screen "0030_Tool Allocation" 1280x800, template "Navigation"
   on GenerateScreen: "ToolAllocation_First"()
   Button "Button_1" at 558,753 size 280x42; TextOff '>>>'
      on Press: function_dd21b452("DB939_Tool_alloc_HMI_AllocList_page", 1); "ToolAllocation_First"()
      Visibility <- "DB939_Tool_alloc_HMI_Limit_allocation_list"
   Button "Button_3" at 326,104 size 451x32; TextOff 'Tool Allocation'
   Button "Button_31" at 872,148 size 242x25; TextOff 'Existing Tools'
   Button "Button_35" at 981,96 size 196x42; TextOff 'TOOL Allocation Automatic'; TextList "Tool_Allocation_Mode"
      ProcessValue <- "DB939_Tool_alloc_HMI_Select_hand_automatic_alloc"
      on Press: InvertBit("DB939_Tool_alloc_HMI_Select_hand_automatic_alloc")
   Button "Button_34" at 167,754 size 280x42; TextOff '<<<'
      on Press: function_b9b71300("DB939_Tool_alloc_HMI_AllocList_page", 1); "ToolAllocation_First"()
      Visibility <- "DB939_Tool_alloc_HMI_AllocList_page"
   Button "b_Decress_ToolAllocation" at 272,104 size 46x32; TextOff 'Text'; PictureOff "left arrow"
      on Click: function_b9b71300("DB939_Tool_alloc_HMI_MH_No_selected", 1); "ToolAllocation_Sec"()
      Visibility <- "DB939_Tool_alloc_HMI_Select_hand_automatic_alloc"
   Button "Button_36" at 432,154 size 34x31; TextOff 'Text'; PictureOff "Tongsampah_1"
      Visibility <- "DB939_Tool_alloc_HMI_Alloc_stationTool{1}"
      on Press: SetTag("DB939_Tool_alloc_HMI_Delete_selected_tool", 1)
   Button "Button_37" at 432,194 size 34x31; TextOff 'Text'; PictureOff "Tongsampah_1"
      Visibility <- "DB939_Tool_alloc_HMI_Alloc_stationTool{2}"
      on Press: SetTag("DB939_Tool_alloc_HMI_Delete_selected_tool", 2)
   Button "Button_38" at 432,234 size 34x31; TextOff 'Text'; PictureOff "Tongsampah_1"
      Visibility <- "DB939_Tool_alloc_HMI_Alloc_stationTool{3}"
      on Press: SetTag("DB939_Tool_alloc_HMI_Delete_selected_tool", 3)
   Button "Button_39" at 432,274 size 34x31; TextOff 'Text'; PictureOff "Tongsampah_1"
      Visibility <- "DB939_Tool_alloc_HMI_Alloc_stationTool{4}"
      on Press: SetTag("DB939_Tool_alloc_HMI_Delete_selected_tool", 4)
   Button "Button_40" at 432,314 size 34x31; TextOff 'Text'; PictureOff "Tongsampah_1"
      Visibility <- "DB939_Tool_alloc_HMI_Alloc_stationTool{5}"
      on Press: SetTag("DB939_Tool_alloc_HMI_Delete_selected_tool", 5)
   Button "Button_41" at 432,354 size 34x31; TextOff 'Text'; PictureOff "Tongsampah_1"
      Visibility <- "DB939_Tool_alloc_HMI_Alloc_stationTool{6}"
      on Press: SetTag("DB939_Tool_alloc_HMI_Delete_selected_tool", 6)
   Button "Button_42" at 432,394 size 34x31; TextOff 'Text'; PictureOff "Tongsampah_1"
      Visibility <- "DB939_Tool_alloc_HMI_Alloc_stationTool{7}"
      on Press: SetTag("DB939_Tool_alloc_HMI_Delete_selected_tool", 7)
   Button "Button_43" at 432,434 size 34x31; TextOff 'Text'; PictureOff "Tongsampah_1"
      Visibility <- "DB939_Tool_alloc_HMI_Alloc_stationTool{8}"
      on Press: SetTag("DB939_Tool_alloc_HMI_Delete_selected_tool", 8)
   Button "Button_44" at 432,474 size 34x31; TextOff 'Text'; PictureOff "Tongsampah_1"
      Visibility <- "DB939_Tool_alloc_HMI_Alloc_stationTool{9}"
      on Press: SetTag("DB939_Tool_alloc_HMI_Delete_selected_tool", 9)
   Button "Button_45" at 432,514 size 34x31; TextOff 'Text'; PictureOff "Tongsampah_1"
      Visibility <- "DB939_Tool_alloc_HMI_Alloc_stationTool{10}"
      on Press: SetTag("DB939_Tool_alloc_HMI_Delete_selected_tool", 10)
   Button "Button_46" at 432,554 size 34x31; TextOff 'Text'; PictureOff "Tongsampah_1"
      Visibility <- "DB939_Tool_alloc_HMI_Alloc_stationTool{11}"
      on Press: SetTag("DB939_Tool_alloc_HMI_Delete_selected_tool", 11)
   Button "Button_47" at 432,594 size 34x31; TextOff 'Text'; PictureOff "Tongsampah_1"
      Visibility <- "DB939_Tool_alloc_HMI_Alloc_stationTool{12}"
      on Press: SetTag("DB939_Tool_alloc_HMI_Delete_selected_tool", 12)
   Button "Button_48" at 432,634 size 34x31; TextOff 'Text'; PictureOff "Tongsampah_1"
      Visibility <- "DB939_Tool_alloc_HMI_Alloc_stationTool{13}"
      on Press: SetTag("DB939_Tool_alloc_HMI_Delete_selected_tool", 13)
   Button "Button_49" at 432,674 size 34x31; TextOff 'Text'; PictureOff "Tongsampah_1"
      Visibility <- "DB939_Tool_alloc_HMI_Alloc_stationTool{14}"
      on Press: SetTag("DB939_Tool_alloc_HMI_Delete_selected_tool", 14)
   Button "Button_50" at 432,714 size 34x31; TextOff 'Text'; PictureOff "Tongsampah_1"
      Visibility <- "DB939_Tool_alloc_HMI_Alloc_stationTool{15}"
      on Press: SetTag("DB939_Tool_alloc_HMI_Delete_selected_tool", 15)
   Button "Button_51" at 807,154 size 34x31; TextOff 'Text'; PictureOff "Tongsampah_1"
      Visibility <- "DB939_Tool_alloc_HMI_Alloc_stationTool{16}"
      on Press: SetTag("DB939_Tool_alloc_HMI_Delete_selected_tool", 16)
   Button "Button_52" at 807,194 size 34x31; TextOff 'Text'; PictureOff "Tongsampah_1"
      Visibility <- "DB939_Tool_alloc_HMI_Alloc_stationTool{17}"
      on Press: SetTag("DB939_Tool_alloc_HMI_Delete_selected_tool", 17)
   Button "Button_53" at 807,234 size 34x31; TextOff 'Text'; PictureOff "Tongsampah_1"
      Visibility <- "DB939_Tool_alloc_HMI_Alloc_stationTool{18}"
      on Press: SetTag("DB939_Tool_alloc_HMI_Delete_selected_tool", 18)
   Button "Button_54" at 807,274 size 34x31; TextOff 'Text'; PictureOff "Tongsampah_1"
      Visibility <- "DB939_Tool_alloc_HMI_Alloc_stationTool{19}"
      on Press: SetTag("DB939_Tool_alloc_HMI_Delete_selected_tool", 19)
   Button "Button_55" at 807,314 size 34x31; TextOff 'Text'; PictureOff "Tongsampah_1"
      Visibility <- "DB939_Tool_alloc_HMI_Alloc_stationTool{20}"
      on Press: SetTag("DB939_Tool_alloc_HMI_Delete_selected_tool", 20)
   Button "Button_56" at 807,354 size 34x31; TextOff 'Text'; PictureOff "Tongsampah_1"
      Visibility <- "DB939_Tool_alloc_HMI_Alloc_stationTool{21}"
      on Press: SetTag("DB939_Tool_alloc_HMI_Delete_selected_tool", 21)
   Button "Button_57" at 807,394 size 34x31; TextOff 'Text'; PictureOff "Tongsampah_1"
      Visibility <- "DB939_Tool_alloc_HMI_Alloc_stationTool{22}"
      on Press: SetTag("DB939_Tool_alloc_HMI_Delete_selected_tool", 22)
   Button "Button_58" at 807,434 size 34x31; TextOff 'Text'; PictureOff "Tongsampah_1"
      Visibility <- "DB939_Tool_alloc_HMI_Alloc_stationTool{23}"
      on Press: SetTag("DB939_Tool_alloc_HMI_Delete_selected_tool", 23)
   Button "Button_59" at 807,474 size 34x31; TextOff 'Text'; PictureOff "Tongsampah_1"
      Visibility <- "DB939_Tool_alloc_HMI_Alloc_stationTool{24}"
      on Press: SetTag("DB939_Tool_alloc_HMI_Delete_selected_tool", 24)
   Button "Button_60" at 807,514 size 34x31; TextOff 'Text'; PictureOff "Tongsampah_1"
      Visibility <- "DB939_Tool_alloc_HMI_Alloc_stationTool{25}"
      on Press: SetTag("DB939_Tool_alloc_HMI_Delete_selected_tool", 25)
   Button "Button_61" at 807,554 size 34x31; TextOff 'Text'; PictureOff "Tongsampah_1"
      Visibility <- "DB939_Tool_alloc_HMI_Alloc_stationTool{26}"
      on Press: SetTag("DB939_Tool_alloc_HMI_Delete_selected_tool", 26)
   Button "Button_62" at 807,594 size 34x31; TextOff 'Text'; PictureOff "Tongsampah_1"
      Visibility <- "DB939_Tool_alloc_HMI_Alloc_stationTool{27}"
      on Press: SetTag("DB939_Tool_alloc_HMI_Delete_selected_tool", 27)
   Button "Button_63" at 807,634 size 34x31; TextOff 'Text'; PictureOff "Tongsampah_1"
      Visibility <- "DB939_Tool_alloc_HMI_Alloc_stationTool{28}"
      on Press: SetTag("DB939_Tool_alloc_HMI_Delete_selected_tool", 28)
   Button "Button_64" at 807,674 size 34x31; TextOff 'Text'; PictureOff "Tongsampah_1"
      Visibility <- "DB939_Tool_alloc_HMI_Alloc_stationTool{29}"
      on Press: SetTag("DB939_Tool_alloc_HMI_Delete_selected_tool", 29)
   Button "Button_65" at 807,714 size 34x31; TextOff 'Text'; PictureOff "Tongsampah_1"
      Visibility <- "DB939_Tool_alloc_HMI_Alloc_stationTool{30}"
      on Press: SetTag("DB939_Tool_alloc_HMI_Delete_selected_tool", 30)
   IOField "I/O field_63" at 971,176 size 144x28; FormatPattern ????????????????????
      ProcessValue <- "DB939_Tool_alloc_HMI_SaveSortProg_name{1}"
      Visibility <- "DB939_Tool_alloc_HMI_SaveSortProgs{1}"
   IOField "I/O field_64" at 971,203 size 144x28; FormatPattern ????????????????????
      ProcessValue <- "DB939_Tool_alloc_HMI_SaveSortProg_name{2}"
      Visibility <- "DB939_Tool_alloc_HMI_SaveSortProgs{2}"
   IOField "I/O field_65" at 971,230 size 144x28; FormatPattern ????????????????????
      ProcessValue <- "DB939_Tool_alloc_HMI_SaveSortProg_name{3}"
      Visibility <- "DB939_Tool_alloc_HMI_SaveSortProgs{3}"
   IOField "I/O field_66" at 971,257 size 144x28; FormatPattern ????????????????????
      ProcessValue <- "DB939_Tool_alloc_HMI_SaveSortProg_name{4}"
      Visibility <- "DB939_Tool_alloc_HMI_SaveSortProgs{4}"
   IOField "I/O field_67" at 971,284 size 144x28; FormatPattern ????????????????????
      ProcessValue <- "DB939_Tool_alloc_HMI_SaveSortProg_name{5}"
      Visibility <- "DB939_Tool_alloc_HMI_SaveSortProgs{5}"
   IOField "I/O field_68" at 971,311 size 144x28; FormatPattern ????????????????????
      ProcessValue <- "DB939_Tool_alloc_HMI_SaveSortProg_name{6}"
      Visibility <- "DB939_Tool_alloc_HMI_SaveSortProgs{6}"
   IOField "I/O field_69" at 971,338 size 144x28; FormatPattern ????????????????????
      ProcessValue <- "DB939_Tool_alloc_HMI_SaveSortProg_name{7}"
      Visibility <- "DB939_Tool_alloc_HMI_SaveSortProgs{7}"
   IOField "I/O field_70" at 971,365 size 144x28; FormatPattern ????????????????????
      ProcessValue <- "DB939_Tool_alloc_HMI_SaveSortProg_name{8}"
      Visibility <- "DB939_Tool_alloc_HMI_SaveSortProgs{8}"
   IOField "I/O field_71" at 971,392 size 144x28; FormatPattern ????????????????????
      ProcessValue <- "DB939_Tool_alloc_HMI_SaveSortProg_name{9}"
      Visibility <- "DB939_Tool_alloc_HMI_SaveSortProgs{9}"
   IOField "I/O field_72" at 971,419 size 144x28; FormatPattern ????????????????????
      ProcessValue <- "DB939_Tool_alloc_HMI_SaveSortProg_name{10}"
      Visibility <- "DB939_Tool_alloc_HMI_SaveSortProgs{10}"
   IOField "I/O field_73" at 971,446 size 144x28; FormatPattern ????????????????????
      ProcessValue <- "DB939_Tool_alloc_HMI_SaveSortProg_name{11}"
      Visibility <- "DB939_Tool_alloc_HMI_SaveSortProgs{11}"
   IOField "I/O field_74" at 971,473 size 144x28; FormatPattern ????????????????????
      ProcessValue <- "DB939_Tool_alloc_HMI_SaveSortProg_name{12}"
      Visibility <- "DB939_Tool_alloc_HMI_SaveSortProgs{12}"
   IOField "I/O field_75" at 971,500 size 144x28; FormatPattern ????????????????????
      ProcessValue <- "DB939_Tool_alloc_HMI_SaveSortProg_name{13}"
      Visibility <- "DB939_Tool_alloc_HMI_SaveSortProgs{13}"
   IOField "I/O field_76" at 971,527 size 144x28; FormatPattern ????????????????????
      ProcessValue <- "DB939_Tool_alloc_HMI_SaveSortProg_name{14}"
      Visibility <- "DB939_Tool_alloc_HMI_SaveSortProgs{14}"
   IOField "I/O field_77" at 971,554 size 144x28; FormatPattern ????????????????????
      ProcessValue <- "DB939_Tool_alloc_HMI_SaveSortProg_name{15}"
      Visibility <- "DB939_Tool_alloc_HMI_SaveSortProgs{15}"
   IOField "I/O field_78" at 971,581 size 144x28; FormatPattern ????????????????????
      ProcessValue <- "DB939_Tool_alloc_HMI_SaveSortProg_name{16}"
      Visibility <- "DB939_Tool_alloc_HMI_SaveSortProgs{16}"
   IOField "I/O field_79" at 971,608 size 144x28; FormatPattern ????????????????????
      ProcessValue <- "DB939_Tool_alloc_HMI_SaveSortProg_name{17}"
      Visibility <- "DB939_Tool_alloc_HMI_SaveSortProgs{17}"
   IOField "I/O field_80" at 971,635 size 144x28; FormatPattern ????????????????????
      ProcessValue <- "DB939_Tool_alloc_HMI_SaveSortProg_name{18}"
      Visibility <- "DB939_Tool_alloc_HMI_SaveSortProgs{18}"
   IOField "I/O field_81" at 971,662 size 144x28; FormatPattern ????????????????????
      ProcessValue <- "DB939_Tool_alloc_HMI_SaveSortProg_name{19}"
      Visibility <- "DB939_Tool_alloc_HMI_SaveSortProgs{19}"
   IOField "I/O field_82" at 971,689 size 144x28; FormatPattern ????????????????????
      ProcessValue <- "DB939_Tool_alloc_HMI_SaveSortProg_name{20}"
      Visibility <- "DB939_Tool_alloc_HMI_SaveSortProgs{20}"
   IOField "I/O field_83" at 877,176 size 96x28; FormatPattern 9999
      ProcessValue <- "DB939_Tool_alloc_HMI_SaveSortProgs{1}"
      Visibility <- "DB939_Tool_alloc_HMI_SaveSortProgs{1}"
   IOField "I/O field_84" at 877,203 size 96x28; FormatPattern 9999
      ProcessValue <- "DB939_Tool_alloc_HMI_SaveSortProgs{2}"
      Visibility <- "DB939_Tool_alloc_HMI_SaveSortProgs{2}"
   IOField "I/O field_85" at 877,230 size 96x28; FormatPattern 9999
      ProcessValue <- "DB939_Tool_alloc_HMI_SaveSortProgs{3}"
      Visibility <- "DB939_Tool_alloc_HMI_SaveSortProgs{3}"
   IOField "I/O field_86" at 877,257 size 96x28; FormatPattern 9999
      ProcessValue <- "DB939_Tool_alloc_HMI_SaveSortProgs{4}"
      Visibility <- "DB939_Tool_alloc_HMI_SaveSortProgs{4}"
   IOField "I/O field_87" at 877,284 size 96x28; FormatPattern 9999
      ProcessValue <- "DB939_Tool_alloc_HMI_SaveSortProgs{5}"
      Visibility <- "DB939_Tool_alloc_HMI_SaveSortProgs{5}"
   IOField "I/O field_88" at 877,311 size 96x28; FormatPattern 9999
      ProcessValue <- "DB939_Tool_alloc_HMI_SaveSortProgs{6}"
      Visibility <- "DB939_Tool_alloc_HMI_SaveSortProgs{6}"
   IOField "I/O field_89" at 877,338 size 96x28; FormatPattern 9999
      ProcessValue <- "DB939_Tool_alloc_HMI_SaveSortProgs{7}"
      Visibility <- "DB939_Tool_alloc_HMI_SaveSortProgs{7}"
   IOField "I/O field_90" at 877,365 size 96x28; FormatPattern 9999
      ProcessValue <- "DB939_Tool_alloc_HMI_SaveSortProgs{8}"
      Visibility <- "DB939_Tool_alloc_HMI_SaveSortProgs{8}"
   IOField "I/O field_91" at 877,392 size 96x28; FormatPattern 9999
      ProcessValue <- "DB939_Tool_alloc_HMI_SaveSortProgs{9}"
      Visibility <- "DB939_Tool_alloc_HMI_SaveSortProgs{9}"
   IOField "I/O field_92" at 877,419 size 96x28; FormatPattern 9999
      ProcessValue <- "DB939_Tool_alloc_HMI_SaveSortProgs{10}"
      Visibility <- "DB939_Tool_alloc_HMI_SaveSortProgs{10}"
   IOField "I/O field_93" at 877,446 size 96x28; FormatPattern 9999
      ProcessValue <- "DB939_Tool_alloc_HMI_SaveSortProgs{11}"
      Visibility <- "DB939_Tool_alloc_HMI_SaveSortProgs{11}"
   IOField "I/O field_94" at 877,473 size 96x28; FormatPattern 9999
      ProcessValue <- "DB939_Tool_alloc_HMI_SaveSortProgs{12}"
      Visibility <- "DB939_Tool_alloc_HMI_SaveSortProgs{12}"
   IOField "I/O field_95" at 877,500 size 96x28; FormatPattern 9999
      ProcessValue <- "DB939_Tool_alloc_HMI_SaveSortProgs{13}"
      Visibility <- "DB939_Tool_alloc_HMI_SaveSortProgs{13}"
   IOField "I/O field_96" at 877,527 size 96x28; FormatPattern 9999
      ProcessValue <- "DB939_Tool_alloc_HMI_SaveSortProgs{14}"
      Visibility <- "DB939_Tool_alloc_HMI_SaveSortProgs{14}"
   IOField "I/O field_97" at 877,554 size 96x28; FormatPattern 9999
      ProcessValue <- "DB939_Tool_alloc_HMI_SaveSortProgs{15}"
      Visibility <- "DB939_Tool_alloc_HMI_SaveSortProgs{15}"
   IOField "I/O field_98" at 877,581 size 96x28; FormatPattern 9999
      ProcessValue <- "DB939_Tool_alloc_HMI_SaveSortProgs{16}"
      Visibility <- "DB939_Tool_alloc_HMI_SaveSortProgs{16}"
   IOField "I/O field_99" at 877,608 size 96x28; FormatPattern 9999
      ProcessValue <- "DB939_Tool_alloc_HMI_SaveSortProgs{17}"
      Visibility <- "DB939_Tool_alloc_HMI_SaveSortProgs{17}"
   IOField "I/O field_100" at 877,635 size 96x28; FormatPattern 9999
      ProcessValue <- "DB939_Tool_alloc_HMI_SaveSortProgs{18}"
      Visibility <- "DB939_Tool_alloc_HMI_SaveSortProgs{18}"
   IOField "I/O field_101" at 877,662 size 96x28; FormatPattern 9999
      ProcessValue <- "DB939_Tool_alloc_HMI_SaveSortProgs{19}"
      Visibility <- "DB939_Tool_alloc_HMI_SaveSortProgs{19}"
   IOField "I/O field_102" at 877,689 size 96x28; FormatPattern 9999
      ProcessValue <- "DB939_Tool_alloc_HMI_SaveSortProgs{20}"
      Visibility <- "DB939_Tool_alloc_HMI_SaveSortProgs{20}"
   Button "Button_66" at 1128,183 size 42x224; TextOff '˄˄˄'
      on Press: SetBit("DB939_Tool_alloc_HMI_SavedProgs_increase")
      Visibility <- "DB939_Tool_alloc_HMI_SavedProgs_increase_visible"
   Button "Button_67" at 1128,485 size 42x224; TextOff 'VVV'
      on Press: SetBit("DB939_Tool_alloc_HMI_SavedProgs_decrease")
      Visibility <- "DB939_Tool_alloc_HMI_SavedProgs_decrease_visible"
   Button "b_Incress_ToolAllocation" at 786,104 size 46x32; TextOff 'Text'; PictureOff "right arrow"
      on Click: function_dd21b452("DB939_Tool_alloc_HMI_MH_No_selected", 1); "ToolAllocation_Sec"()
      Visibility <- "DB939_Tool_alloc_HMI_Select_hand_automatic_alloc"
   IOField "I/O field_5" at 179,152 size 73x35; Authorization "User administration"; FormatPattern 999
      ProcessValue <- "DB939_Tool_alloc_HMI_Alloc_stationTool{1}"
      Visibility <- "DB939_Tool_alloc_HMI_Limit_allocation_list"
      Appearance <- "DB939_Tool_alloc_HMI_Selected_prog"
   Button "Button_6" at 123,152 size 50x35; TextOff '.'
      Visibility <- "DB939_Tool_alloc_HMI_Limit_allocation_list"
      on Press: SetTag("DB939_Tool_alloc_HMI_Selected_prog", 1)
      Appearance <- "DB939_Tool_alloc_HMI_Selected_prog"
   Button "Button_2" at 123,192 size 50x35; TextOff '.'
      Visibility <- "DB939_Tool_alloc_HMI_Limit_allocation_list"
      on Press: SetTag("DB939_Tool_alloc_HMI_Selected_prog", 2)
      Appearance <- "DB939_Tool_alloc_HMI_Selected_prog"
   Button "Button_4" at 123,232 size 50x35; TextOff '.'
      Visibility <- "DB939_Tool_alloc_HMI_Limit_allocation_list"
      on Press: SetTag("DB939_Tool_alloc_HMI_Selected_prog", 3)
      Appearance <- "DB939_Tool_alloc_HMI_Selected_prog"
   Button "Button_5" at 123,272 size 50x35; TextOff '.'
      Visibility <- "DB939_Tool_alloc_HMI_Limit_allocation_list"
      on Press: SetTag("DB939_Tool_alloc_HMI_Selected_prog", 4)
      Appearance <- "DB939_Tool_alloc_HMI_Selected_prog"
   Button "Button_7" at 123,312 size 50x35; TextOff '.'
      Visibility <- "DB939_Tool_alloc_HMI_Limit_allocation_list"
      on Press: SetTag("DB939_Tool_alloc_HMI_Selected_prog", 5)
      Appearance <- "DB939_Tool_alloc_HMI_Selected_prog"
   Button "Button_8" at 123,352 size 50x35; TextOff '.'
      Visibility <- "DB939_Tool_alloc_HMI_Limit_allocation_list"
      on Press: SetTag("DB939_Tool_alloc_HMI_Selected_prog", 6)
      Appearance <- "DB939_Tool_alloc_HMI_Selected_prog"
   Button "Button_9" at 123,392 size 50x35; TextOff '.'
      Visibility <- "DB939_Tool_alloc_HMI_Limit_allocation_list"
      on Press: SetTag("DB939_Tool_alloc_HMI_Selected_prog", 7)
      Appearance <- "DB939_Tool_alloc_HMI_Selected_prog"
   Button "Button_10" at 123,432 size 50x35; TextOff '.'
      on Press: SetTag("DB939_Tool_alloc_HMI_Selected_prog", 8)
      Appearance <- "DB939_Tool_alloc_HMI_Selected_prog"
      Visibility <- "DB939_Tool_alloc_HMI_Limit_allocation_list"
   Button "Button_11" at 123,472 size 50x35; TextOff '.'
      Visibility <- "DB939_Tool_alloc_HMI_Limit_allocation_list"
      on Press: SetTag("DB939_Tool_alloc_HMI_Selected_prog", 9)
      Appearance <- "DB939_Tool_alloc_HMI_Selected_prog"
   Button "Button_12" at 123,512 size 50x35; TextOff '.'
      Visibility <- "DB939_Tool_alloc_HMI_Limit_allocation_list"
      on Press: SetTag("DB939_Tool_alloc_HMI_Selected_prog", 10)
      Appearance <- "DB939_Tool_alloc_HMI_Selected_prog"
   Button "Button_13" at 123,552 size 50x35; TextOff '.'
      Visibility <- "DB939_Tool_alloc_HMI_Limit_allocation_list"
      on Press: SetTag("DB939_Tool_alloc_HMI_Selected_prog", 11)
      Appearance <- "DB939_Tool_alloc_HMI_Selected_prog"
   Button "Button_14" at 123,592 size 50x35; TextOff '.'
      Visibility <- "DB939_Tool_alloc_HMI_Limit_allocation_list"
      on Press: SetTag("DB939_Tool_alloc_HMI_Selected_prog", 12)
      Appearance <- "DB939_Tool_alloc_HMI_Selected_prog"
   Button "Button_15" at 123,632 size 50x35; TextOff '.'
      Visibility <- "DB939_Tool_alloc_HMI_Limit_allocation_list"
      on Press: SetTag("DB939_Tool_alloc_HMI_Selected_prog", 13)
      Appearance <- "DB939_Tool_alloc_HMI_Selected_prog"
   Button "Button_16" at 123,672 size 50x35; TextOff '.'
      Visibility <- "DB939_Tool_alloc_HMI_Limit_allocation_list"
      on Press: SetTag("DB939_Tool_alloc_HMI_Selected_prog", 14)
      Appearance <- "DB939_Tool_alloc_HMI_Selected_prog"
   Button "Button_17" at 496,152 size 50x35; TextOff '.'
      Visibility <- "DB939_Tool_alloc_HMI_Limit_allocation_list"
      on Press: SetTag("DB939_Tool_alloc_HMI_Selected_prog", 16)
      Appearance <- "DB939_Tool_alloc_HMI_Selected_prog"
   Button "Button_18" at 496,192 size 50x35; TextOff '.'
      Visibility <- "DB939_Tool_alloc_HMI_Limit_allocation_list"
      on Press: SetTag("DB939_Tool_alloc_HMI_Selected_prog", 17)
      Appearance <- "DB939_Tool_alloc_HMI_Selected_prog"
   Button "Button_19" at 496,232 size 50x35; TextOff '.'
      Visibility <- "DB939_Tool_alloc_HMI_Limit_allocation_list"
      on Press: SetTag("DB939_Tool_alloc_HMI_Selected_prog", 18)
      Appearance <- "DB939_Tool_alloc_HMI_Selected_prog"
   Button "Button_20" at 496,272 size 50x35; TextOff '.'
      Visibility <- "DB939_Tool_alloc_HMI_Limit_allocation_list"
      on Press: SetTag("DB939_Tool_alloc_HMI_Selected_prog", 19)
      Appearance <- "DB939_Tool_alloc_HMI_Selected_prog"
   Button "Button_21" at 496,312 size 50x35; TextOff '.'
      Visibility <- "DB939_Tool_alloc_HMI_Limit_allocation_list"
      on Press: SetTag("DB939_Tool_alloc_HMI_Selected_prog", 20)
      Appearance <- "DB939_Tool_alloc_HMI_Selected_prog"
   Button "Button_22" at 496,352 size 50x35; TextOff '.'
      Visibility <- "DB939_Tool_alloc_HMI_Limit_allocation_list"
      on Press: SetTag("DB939_Tool_alloc_HMI_Selected_prog", 21)
      Appearance <- "DB939_Tool_alloc_HMI_Selected_prog"
   Button "Button_23" at 496,392 size 50x35; TextOff '.'
      Visibility <- "DB939_Tool_alloc_HMI_Limit_allocation_list"
      on Press: SetTag("DB939_Tool_alloc_HMI_Selected_prog", 22)
      Appearance <- "DB939_Tool_alloc_HMI_Selected_prog"
   Button "Button_24" at 496,432 size 50x35; TextOff '.'
      Visibility <- "DB939_Tool_alloc_HMI_Limit_allocation_list"
      on Press: SetTag("DB939_Tool_alloc_HMI_Selected_prog", 23)
      Appearance <- "DB939_Tool_alloc_HMI_Selected_prog"
   Button "Button_25" at 496,472 size 50x35; TextOff 'Text'
      Visibility <- "DB939_Tool_alloc_HMI_Limit_allocation_list"
      on Press: SetTag("DB939_Tool_alloc_HMI_Selected_prog", 24)
      Appearance <- "DB939_Tool_alloc_HMI_Selected_prog"
   Button "Button_26" at 496,512 size 50x35; TextOff 'Text'
      Visibility <- "DB939_Tool_alloc_HMI_Limit_allocation_list"
      on Press: SetTag("DB939_Tool_alloc_HMI_Selected_prog", 25)
      Appearance <- "DB939_Tool_alloc_HMI_Selected_prog"
   Button "Button_27" at 496,552 size 50x35; TextOff '.'
      Visibility <- "DB939_Tool_alloc_HMI_Limit_allocation_list"
      on Press: SetTag("DB939_Tool_alloc_HMI_Selected_prog", 26)
      Appearance <- "DB939_Tool_alloc_HMI_Selected_prog"
   Button "Button_28" at 496,592 size 50x35; TextOff '.'
      Visibility <- "DB939_Tool_alloc_HMI_Limit_allocation_list"
      on Press: SetTag("DB939_Tool_alloc_HMI_Selected_prog", 27)
      Appearance <- "DB939_Tool_alloc_HMI_Selected_prog"
   Button "Button_29" at 496,632 size 50x35; TextOff '.'
      Visibility <- "DB939_Tool_alloc_HMI_Limit_allocation_list"
      on Press: SetTag("DB939_Tool_alloc_HMI_Selected_prog", 28)
      Appearance <- "DB939_Tool_alloc_HMI_Selected_prog"
   Button "Button_30" at 496,672 size 50x35; TextOff '.'
      Visibility <- "DB939_Tool_alloc_HMI_Limit_allocation_list"
      on Press: SetTag("DB939_Tool_alloc_HMI_Selected_prog", 29)
      Appearance <- "DB939_Tool_alloc_HMI_Selected_prog"
   IOField "Station_Tool_2" at 179,192 size 73x35; Authorization "User administration"; FormatPattern 999
      ProcessValue <- "DB939_Tool_alloc_HMI_Alloc_stationTool{2}"
      Visibility <- "DB939_Tool_alloc_HMI_Limit_allocation_list"
      Appearance <- "DB939_Tool_alloc_HMI_Selected_prog"
   IOField "I/O field_2" at 179,232 size 73x35; Authorization "User administration"; FormatPattern 999
      ProcessValue <- "DB939_Tool_alloc_HMI_Alloc_stationTool{3}"
      Visibility <- "DB939_Tool_alloc_HMI_Limit_allocation_list"
      Appearance <- "DB939_Tool_alloc_HMI_Selected_prog"
   IOField "I/O field_3" at 179,272 size 73x35; Authorization "User administration"; FormatPattern 999
      ProcessValue <- "DB939_Tool_alloc_HMI_Alloc_stationTool{4}"
      Visibility <- "DB939_Tool_alloc_HMI_Limit_allocation_list"
      Appearance <- "DB939_Tool_alloc_HMI_Selected_prog"
   IOField "I/O field_4" at 179,312 size 73x35; Authorization "User administration"; FormatPattern 999
      ProcessValue <- "DB939_Tool_alloc_HMI_Alloc_stationTool{5}"
      Visibility <- "DB939_Tool_alloc_HMI_Limit_allocation_list"
      Appearance <- "DB939_Tool_alloc_HMI_Selected_prog"
   IOField "I/O field_6" at 179,352 size 73x35; Authorization "User administration"; FormatPattern 999
      ProcessValue <- "DB939_Tool_alloc_HMI_Alloc_stationTool{6}"
      Visibility <- "DB939_Tool_alloc_HMI_Limit_allocation_list"
      Appearance <- "DB939_Tool_alloc_HMI_Selected_prog"
   IOField "I/O field_7" at 179,392 size 73x35; Authorization "User administration"; FormatPattern 999
      ProcessValue <- "DB939_Tool_alloc_HMI_Alloc_stationTool{7}"
      Visibility <- "DB939_Tool_alloc_HMI_Limit_allocation_list"
      Appearance <- "DB939_Tool_alloc_HMI_Selected_prog"
   IOField "I/O field_8" at 179,432 size 73x35; Authorization "User administration"; FormatPattern 999
      ProcessValue <- "DB939_Tool_alloc_HMI_Alloc_stationTool{8}"
      Appearance <- "DB939_Tool_alloc_HMI_Selected_prog"
      Visibility <- "DB939_Tool_alloc_HMI_Limit_allocation_list"
   IOField "I/O field_9" at 179,472 size 73x35; Authorization "User administration"; FormatPattern 999
      ProcessValue <- "DB939_Tool_alloc_HMI_Alloc_stationTool{9}"
      Visibility <- "DB939_Tool_alloc_HMI_Limit_allocation_list"
      Appearance <- "DB939_Tool_alloc_HMI_Selected_prog"
   IOField "I/O field_10" at 179,512 size 73x35; Authorization "User administration"; FormatPattern 999
      ProcessValue <- "DB939_Tool_alloc_HMI_Alloc_stationTool{10}"
      Visibility <- "DB939_Tool_alloc_HMI_Limit_allocation_list"
      Appearance <- "DB939_Tool_alloc_HMI_Selected_prog"
   IOField "I/O field_11" at 179,552 size 73x35; Authorization "User administration"; FormatPattern 999
      ProcessValue <- "DB939_Tool_alloc_HMI_Alloc_stationTool{11}"
      Visibility <- "DB939_Tool_alloc_HMI_Limit_allocation_list"
      Appearance <- "DB939_Tool_alloc_HMI_Selected_prog"
   IOField "I/O field_12" at 179,592 size 73x35; Authorization "User administration"; FormatPattern 999
      ProcessValue <- "DB939_Tool_alloc_HMI_Alloc_stationTool{12}"
      Visibility <- "DB939_Tool_alloc_HMI_Limit_allocation_list"
      Appearance <- "DB939_Tool_alloc_HMI_Selected_prog"
   IOField "I/O field_13" at 179,632 size 73x35; Authorization "User administration"; FormatPattern 999
      ProcessValue <- "DB939_Tool_alloc_HMI_Alloc_stationTool{13}"
      Visibility <- "DB939_Tool_alloc_HMI_Limit_allocation_list"
      Appearance <- "DB939_Tool_alloc_HMI_Selected_prog"
   IOField "I/O field_14" at 179,672 size 73x35; Authorization "User administration"; FormatPattern 999
      ProcessValue <- "DB939_Tool_alloc_HMI_Alloc_stationTool{14}"
      Visibility <- "DB939_Tool_alloc_HMI_Limit_allocation_list"
      Appearance <- "DB939_Tool_alloc_HMI_Selected_prog"
   IOField "I/O field_15" at 552,152 size 73x35; Authorization "User administration"; FormatPattern 999
      ProcessValue <- "DB939_Tool_alloc_HMI_Alloc_stationTool{16}"
      Visibility <- "DB939_Tool_alloc_HMI_Limit_allocation_list"
      Appearance <- "DB939_Tool_alloc_HMI_Selected_prog"
   IOField "I/O field_16" at 552,192 size 73x35; Authorization "User administration"; FormatPattern 999
      ProcessValue <- "DB939_Tool_alloc_HMI_Alloc_stationTool{17}"
      Visibility <- "DB939_Tool_alloc_HMI_Limit_allocation_list"
      Appearance <- "DB939_Tool_alloc_HMI_Selected_prog"
   IOField "I/O field_17" at 552,232 size 73x35; Authorization "User administration"; FormatPattern 999
      ProcessValue <- "DB939_Tool_alloc_HMI_Alloc_stationTool{18}"
      Visibility <- "DB939_Tool_alloc_HMI_Limit_allocation_list"
      Appearance <- "DB939_Tool_alloc_HMI_Selected_prog"
   IOField "I/O field_18" at 552,272 size 73x35; Authorization "User administration"; FormatPattern 999
      ProcessValue <- "DB939_Tool_alloc_HMI_Alloc_stationTool{19}"
      Visibility <- "DB939_Tool_alloc_HMI_Limit_allocation_list"
      Appearance <- "DB939_Tool_alloc_HMI_Selected_prog"
   IOField "I/O field_19" at 552,312 size 73x35; Authorization "User administration"; FormatPattern 999
      ProcessValue <- "DB939_Tool_alloc_HMI_Alloc_stationTool{20}"
      Visibility <- "DB939_Tool_alloc_HMI_Limit_allocation_list"
      Appearance <- "DB939_Tool_alloc_HMI_Selected_prog"
   IOField "I/O field_20" at 552,352 size 73x35; Authorization "User administration"; FormatPattern 999
      ProcessValue <- "DB939_Tool_alloc_HMI_Alloc_stationTool{21}"
      Visibility <- "DB939_Tool_alloc_HMI_Limit_allocation_list"
      Appearance <- "DB939_Tool_alloc_HMI_Selected_prog"
   IOField "I/O field_21" at 552,392 size 73x35; Authorization "User administration"; FormatPattern 999
      ProcessValue <- "DB939_Tool_alloc_HMI_Alloc_stationTool{22}"
      Visibility <- "DB939_Tool_alloc_HMI_Limit_allocation_list"
      Appearance <- "DB939_Tool_alloc_HMI_Selected_prog"
   IOField "I/O field_22" at 552,432 size 73x35; Authorization "User administration"; FormatPattern 999
      ProcessValue <- "DB939_Tool_alloc_HMI_Alloc_stationTool{23}"
      Visibility <- "DB939_Tool_alloc_HMI_Limit_allocation_list"
      Appearance <- "DB939_Tool_alloc_HMI_Selected_prog"
   IOField "I/O field_23" at 552,472 size 73x35; Authorization "User administration"; FormatPattern 999
      ProcessValue <- "DB939_Tool_alloc_HMI_Alloc_stationTool{24}"
      Visibility <- "DB939_Tool_alloc_HMI_Limit_allocation_list"
      Appearance <- "DB939_Tool_alloc_HMI_Selected_prog"
   IOField "I/O field_24" at 552,512 size 73x35; Authorization "User administration"; FormatPattern 999
      ProcessValue <- "DB939_Tool_alloc_HMI_Alloc_stationTool{25}"
      Visibility <- "DB939_Tool_alloc_HMI_Limit_allocation_list"
      Appearance <- "DB939_Tool_alloc_HMI_Selected_prog"
   IOField "I/O field_25" at 552,552 size 73x35; Authorization "User administration"; FormatPattern 999
      ProcessValue <- "DB939_Tool_alloc_HMI_Alloc_stationTool{26}"
      Visibility <- "DB939_Tool_alloc_HMI_Limit_allocation_list"
      Appearance <- "DB939_Tool_alloc_HMI_Selected_prog"
   IOField "I/O field_26" at 552,592 size 73x35; Authorization "User administration"; FormatPattern 999
      ProcessValue <- "DB939_Tool_alloc_HMI_Alloc_stationTool{27}"
      Visibility <- "DB939_Tool_alloc_HMI_Limit_allocation_list"
      Appearance <- "DB939_Tool_alloc_HMI_Selected_prog"
   IOField "I/O field_27" at 552,632 size 73x35; Authorization "User administration"; FormatPattern 999
      ProcessValue <- "DB939_Tool_alloc_HMI_Alloc_stationTool{28}"
      Visibility <- "DB939_Tool_alloc_HMI_Limit_allocation_list"
      Appearance <- "DB939_Tool_alloc_HMI_Selected_prog"
   IOField "I/O field_28" at 552,672 size 73x35; Authorization "User administration"; FormatPattern 999
      ProcessValue <- "DB939_Tool_alloc_HMI_Alloc_stationTool{29}"
      Visibility <- "DB939_Tool_alloc_HMI_Limit_allocation_list"
      Appearance <- "DB939_Tool_alloc_HMI_Selected_prog"
   IOField "I/O field_29" at 259,152 size 159x35; Authorization "User administration"; FormatPattern ????????????????????
      ProcessValue <- "DB939_Tool_alloc_HMI_Alloc_tool_name{1}"
      Visibility <- "DB939_Tool_alloc_HMI_Limit_allocation_list"
      Appearance <- "DB939_Tool_alloc_HMI_Selected_prog"
   IOField "I/O field_30" at 260,192 size 159x35; Authorization "User administration"; FormatPattern ????????????????????
      ProcessValue <- "DB939_Tool_alloc_HMI_Alloc_tool_name{2}"
      Visibility <- "DB939_Tool_alloc_HMI_Limit_allocation_list"
      Appearance <- "DB939_Tool_alloc_HMI_Selected_prog"
   IOField "I/O field_31" at 260,232 size 159x35; Authorization "User administration"; FormatPattern ????????????????????
      ProcessValue <- "DB939_Tool_alloc_HMI_Alloc_tool_name{3}"
      Visibility <- "DB939_Tool_alloc_HMI_Limit_allocation_list"
      Appearance <- "DB939_Tool_alloc_HMI_Selected_prog"
   IOField "I/O field_32" at 260,272 size 159x35; Authorization "User administration"; FormatPattern ????????????????????
      ProcessValue <- "DB939_Tool_alloc_HMI_Alloc_tool_name{4}"
      Visibility <- "DB939_Tool_alloc_HMI_Limit_allocation_list"
      Appearance <- "DB939_Tool_alloc_HMI_Selected_prog"
   IOField "I/O field_33" at 260,312 size 159x35; Authorization "User administration"; FormatPattern ????????????????????
      ProcessValue <- "DB939_Tool_alloc_HMI_Alloc_tool_name{5}"
      Visibility <- "DB939_Tool_alloc_HMI_Limit_allocation_list"
      Appearance <- "DB939_Tool_alloc_HMI_Selected_prog"
   IOField "I/O field_34" at 260,352 size 159x35; Authorization "User administration"; FormatPattern ????????????????????
      ProcessValue <- "DB939_Tool_alloc_HMI_Alloc_tool_name{6}"
      Visibility <- "DB939_Tool_alloc_HMI_Limit_allocation_list"
      Appearance <- "DB939_Tool_alloc_HMI_Selected_prog"
   IOField "I/O field_35" at 260,392 size 159x35; Authorization "User administration"; FormatPattern ????????????????????
      ProcessValue <- "DB939_Tool_alloc_HMI_Alloc_tool_name{7}"
      Visibility <- "DB939_Tool_alloc_HMI_Limit_allocation_list"
      Appearance <- "DB939_Tool_alloc_HMI_Selected_prog"
   IOField "I/O field_36" at 260,432 size 159x35; Authorization "User administration"; FormatPattern ????????????????????
      ProcessValue <- "DB939_Tool_alloc_HMI_Alloc_tool_name{8}"
      Appearance <- "DB939_Tool_alloc_HMI_Selected_prog"
      Visibility <- "DB939_Tool_alloc_HMI_Limit_allocation_list"
   IOField "I/O field_37" at 260,472 size 159x35; Authorization "User administration"; FormatPattern ????????????????????
      ProcessValue <- "DB939_Tool_alloc_HMI_Alloc_tool_name{9}"
      Visibility <- "DB939_Tool_alloc_HMI_Limit_allocation_list"
      Appearance <- "DB939_Tool_alloc_HMI_Selected_prog"
   IOField "I/O field_38" at 260,512 size 159x35; Authorization "User administration"; FormatPattern ????????????????????
      ProcessValue <- "DB939_Tool_alloc_HMI_Alloc_tool_name{10}"
      Visibility <- "DB939_Tool_alloc_HMI_Limit_allocation_list"
      Appearance <- "DB939_Tool_alloc_HMI_Selected_prog"
   IOField "I/O field_39" at 260,552 size 159x35; Authorization "User administration"; FormatPattern ????????????????????
      ProcessValue <- "DB939_Tool_alloc_HMI_Alloc_tool_name{11}"
      Visibility <- "DB939_Tool_alloc_HMI_Limit_allocation_list"
      Appearance <- "DB939_Tool_alloc_HMI_Selected_prog"
   IOField "I/O field_40" at 260,592 size 159x35; Authorization "User administration"; FormatPattern ????????????????????
      ProcessValue <- "DB939_Tool_alloc_HMI_Alloc_tool_name{12}"
      Visibility <- "DB939_Tool_alloc_HMI_Limit_allocation_list"
      Appearance <- "DB939_Tool_alloc_HMI_Selected_prog"
   IOField "I/O field_41" at 260,632 size 159x35; Authorization "User administration"; FormatPattern ????????????????????
      ProcessValue <- "DB939_Tool_alloc_HMI_Alloc_tool_name{13}"
      Visibility <- "DB939_Tool_alloc_HMI_Limit_allocation_list"
      Appearance <- "DB939_Tool_alloc_HMI_Selected_prog"
   IOField "I/O field_42" at 260,672 size 159x35; Authorization "User administration"; FormatPattern ????????????????????
      ProcessValue <- "DB939_Tool_alloc_HMI_Alloc_tool_name{14}"
      Visibility <- "DB939_Tool_alloc_HMI_Limit_allocation_list"
      Appearance <- "DB939_Tool_alloc_HMI_Selected_prog"
   IOField "I/O field_43" at 632,152 size 159x35; Authorization "User administration"; FormatPattern ????????????????????
      ProcessValue <- "DB939_Tool_alloc_HMI_Alloc_tool_name{16}"
      Visibility <- "DB939_Tool_alloc_HMI_Limit_allocation_list"
      Appearance <- "DB939_Tool_alloc_HMI_Selected_prog"
   IOField "I/O field_44" at 632,192 size 159x35; Authorization "User administration"; FormatPattern ????????????????????
      ProcessValue <- "DB939_Tool_alloc_HMI_Alloc_tool_name{17}"
      Visibility <- "DB939_Tool_alloc_HMI_Limit_allocation_list"
      Appearance <- "DB939_Tool_alloc_HMI_Selected_prog"
   IOField "I/O field_45" at 632,232 size 159x35; Authorization "User administration"; FormatPattern ????????????????????
      ProcessValue <- "DB939_Tool_alloc_HMI_Alloc_tool_name{18}"
      Visibility <- "DB939_Tool_alloc_HMI_Limit_allocation_list"
      Appearance <- "DB939_Tool_alloc_HMI_Selected_prog"
   IOField "I/O field_46" at 632,272 size 159x35; Authorization "User administration"; FormatPattern ????????????????????
      ProcessValue <- "DB939_Tool_alloc_HMI_Alloc_tool_name{19}"
      Visibility <- "DB939_Tool_alloc_HMI_Limit_allocation_list"
      Appearance <- "DB939_Tool_alloc_HMI_Selected_prog"
   IOField "I/O field_47" at 632,312 size 159x35; Authorization "User administration"; FormatPattern ????????????????????
      ProcessValue <- "DB939_Tool_alloc_HMI_Alloc_tool_name{20}"
      Visibility <- "DB939_Tool_alloc_HMI_Limit_allocation_list"
      Appearance <- "DB939_Tool_alloc_HMI_Selected_prog"
   IOField "I/O field_48" at 632,352 size 159x35; Authorization "User administration"; FormatPattern ????????????????????
      ProcessValue <- "DB939_Tool_alloc_HMI_Alloc_tool_name{21}"
      Visibility <- "DB939_Tool_alloc_HMI_Limit_allocation_list"
      Appearance <- "DB939_Tool_alloc_HMI_Selected_prog"
   IOField "I/O field_49" at 632,392 size 159x35; Authorization "User administration"; FormatPattern ????????????????????
      ProcessValue <- "DB939_Tool_alloc_HMI_Alloc_tool_name{22}"
      Visibility <- "DB939_Tool_alloc_HMI_Limit_allocation_list"
      Appearance <- "DB939_Tool_alloc_HMI_Selected_prog"
   IOField "I/O field_50" at 632,432 size 159x35; Authorization "User administration"; FormatPattern ????????????????????
      ProcessValue <- "DB939_Tool_alloc_HMI_Alloc_tool_name{23}"
      Visibility <- "DB939_Tool_alloc_HMI_Limit_allocation_list"
      Appearance <- "DB939_Tool_alloc_HMI_Selected_prog"
   IOField "I/O field_51" at 632,472 size 159x35; Authorization "User administration"; FormatPattern ????????????????????
      ProcessValue <- "DB939_Tool_alloc_HMI_Alloc_tool_name{24}"
      Visibility <- "DB939_Tool_alloc_HMI_Limit_allocation_list"
      Appearance <- "DB939_Tool_alloc_HMI_Selected_prog"
   IOField "I/O field_52" at 632,512 size 159x35; Authorization "User administration"; FormatPattern ????????????????????
      ProcessValue <- "DB939_Tool_alloc_HMI_Alloc_tool_name{25}"
      Visibility <- "DB939_Tool_alloc_HMI_Limit_allocation_list"
      Appearance <- "DB939_Tool_alloc_HMI_Selected_prog"
   IOField "I/O field_53" at 632,552 size 159x35; Authorization "User administration"; FormatPattern ????????????????????
      ProcessValue <- "DB939_Tool_alloc_HMI_Alloc_tool_name{26}"
      Visibility <- "DB939_Tool_alloc_HMI_Limit_allocation_list"
      Appearance <- "DB939_Tool_alloc_HMI_Selected_prog"
   IOField "I/O field_54" at 632,592 size 159x35; Authorization "User administration"; FormatPattern ????????????????????
      ProcessValue <- "DB939_Tool_alloc_HMI_Alloc_tool_name{27}"
      Visibility <- "DB939_Tool_alloc_HMI_Limit_allocation_list"
      Appearance <- "DB939_Tool_alloc_HMI_Selected_prog"
   IOField "I/O field_55" at 632,632 size 159x35; Authorization "User administration"; FormatPattern ????????????????????
      ProcessValue <- "DB939_Tool_alloc_HMI_Alloc_tool_name{28}"
      Visibility <- "DB939_Tool_alloc_HMI_Limit_allocation_list"
      Appearance <- "DB939_Tool_alloc_HMI_Selected_prog"
   IOField "I/O field_56" at 632,672 size 159x35; Authorization "User administration"; FormatPattern ????????????????????
      ProcessValue <- "DB939_Tool_alloc_HMI_Alloc_tool_name{29}"
      Visibility <- "DB939_Tool_alloc_HMI_Limit_allocation_list"
      Appearance <- "DB939_Tool_alloc_HMI_Selected_prog"
   Button "Button_32" at 496,710 size 50x35; TextOff '.'
      Visibility <- "DB939_Tool_alloc_HMI_Limit_allocation_list"
      on Press: SetTag("DB939_Tool_alloc_HMI_Selected_prog", 30)
      Appearance <- "DB939_Tool_alloc_HMI_Selected_prog"
   IOField "I/O field_57" at 551,707 size 73x35; Authorization "User administration"; FormatPattern 999
      ProcessValue <- "DB939_Tool_alloc_HMI_Alloc_stationTool{30}"
      Visibility <- "DB939_Tool_alloc_HMI_Limit_allocation_list"
      Appearance <- "DB939_Tool_alloc_HMI_Selected_prog"
   IOField "I/O field_58" at 631,707 size 159x35; Authorization "User administration"; FormatPattern ????????????????????
      ProcessValue <- "DB939_Tool_alloc_HMI_Alloc_tool_name{30}"
      Visibility <- "DB939_Tool_alloc_HMI_Limit_allocation_list"
      Appearance <- "DB939_Tool_alloc_HMI_Selected_prog"
   Button "Button_33" at 124,713 size 50x35; TextOff '.'
      Visibility <- "DB939_Tool_alloc_HMI_Limit_allocation_list"
      on Press: SetTag("DB939_Tool_alloc_HMI_Selected_prog", 15)
      Appearance <- "DB939_Tool_alloc_HMI_Selected_prog"
   IOField "I/O field_59" at 180,712 size 73x35; Authorization "User administration"; FormatPattern 999
      ProcessValue <- "DB939_Tool_alloc_HMI_Alloc_stationTool{15}"
      Visibility <- "DB939_Tool_alloc_HMI_Limit_allocation_list"
      Appearance <- "DB939_Tool_alloc_HMI_Selected_prog"
   IOField "I/O field_60" at 260,712 size 159x35; Authorization "User administration"; FormatPattern ????????????????????
      ProcessValue <- "DB939_Tool_alloc_HMI_Alloc_tool_name{15}"
      Visibility <- "DB939_Tool_alloc_HMI_Limit_allocation_list"
      Appearance <- "DB939_Tool_alloc_HMI_Selected_prog"
   IOField "I/O field_61" at 465,756 size 73x35; FormatPattern 999
      ProcessValue <- "DB939_Tool_alloc_HMI_AllocList_page"
      Visibility <- "DB939_Tool_alloc_HMI_Limit_allocation_list"
   IOField "I/O field_62" at 734,108 size 39x25; FormatPattern 99
      ProcessValue <- "DB939_Tool_alloc_HMI_MH_No_selected"
      Visibility <- "DB939_Tool_alloc_HMI_Select_hand_automatic_alloc"
   Button "Button_68" at 864,176 size 256x28; TextOff 'Text'
      on Press: SetTag("Tag_1", 1)
      Visibility <- "DB939_Tool_alloc_HMI_SaveSortProgs{1}"
   Button "Button_69" at 864,203 size 256x28; TextOff 'Text'
      on Press: SetTag("Tag_1", 2)
      Visibility <- "DB939_Tool_alloc_HMI_SaveSortProgs{2}"
   Button "Button_70" at 864,230 size 256x28; TextOff 'Text'
      on Press: SetTag("Tag_1", 3)
      Visibility <- "DB939_Tool_alloc_HMI_SaveSortProgs{3}"
   Button "Button_71" at 864,257 size 256x28; TextOff 'Text'
      on Press: SetTag("Tag_1", 4)
      Visibility <- "DB939_Tool_alloc_HMI_SaveSortProgs{4}"
   Button "Button_72" at 864,284 size 256x28; TextOff 'Text'
      on Press: SetTag("Tag_1", 5)
      Visibility <- "DB939_Tool_alloc_HMI_SaveSortProgs{5}"
   Button "Button_73" at 864,311 size 256x28; TextOff 'Text'
      on Press: SetTag("Tag_1", 6)
      Visibility <- "DB939_Tool_alloc_HMI_SaveSortProgs{6}"
   Button "Button_74" at 864,338 size 256x28; TextOff 'Text'
      on Press: SetTag("Tag_1", 7)
      Visibility <- "DB939_Tool_alloc_HMI_SaveSortProgs{7}"
   Button "Button_75" at 864,365 size 256x28; TextOff 'Text'
      on Press: SetTag("Tag_1", 8)
      Visibility <- "DB939_Tool_alloc_HMI_SaveSortProgs{8}"
   Button "Button_76" at 864,392 size 256x28; TextOff 'Text'
      on Press: SetTag("Tag_1", 9)
      Visibility <- "DB939_Tool_alloc_HMI_SaveSortProgs{9}"
   Button "Button_77" at 864,419 size 256x28; TextOff 'Text'
      on Press: SetTag("Tag_1", 10)
      Visibility <- "DB939_Tool_alloc_HMI_SaveSortProgs{10}"
   Button "Button_78" at 864,446 size 256x28; TextOff 'Text'
      on Press: SetTag("Tag_1", 11)
      Visibility <- "DB939_Tool_alloc_HMI_SaveSortProgs{11}"
   Button "Button_79" at 864,473 size 256x28; TextOff 'Text'
      on Press: SetTag("Tag_1", 12)
      Visibility <- "DB939_Tool_alloc_HMI_SaveSortProgs{12}"
   Button "Button_80" at 864,500 size 256x28; TextOff 'Text'
      on Press: SetTag("Tag_1", 13)
      Visibility <- "DB939_Tool_alloc_HMI_SaveSortProgs{13}"
   Button "Button_81" at 864,527 size 256x28; TextOff 'Text'
      on Press: SetTag("Tag_1", 14)
      Visibility <- "DB939_Tool_alloc_HMI_SaveSortProgs{14}"
   Button "Button_82" at 864,554 size 256x28; TextOff 'Text'
      on Press: SetTag("Tag_1", 15)
      Visibility <- "DB939_Tool_alloc_HMI_SaveSortProgs{15}"
   Button "Button_83" at 864,581 size 256x28; TextOff 'Text'
      on Press: SetTag("Tag_1", 16)
      Visibility <- "DB939_Tool_alloc_HMI_SaveSortProgs{16}"
   Button "Button_84" at 864,608 size 256x28; TextOff 'Text'
      on Press: SetTag("Tag_1", 17)
      Visibility <- "DB939_Tool_alloc_HMI_SaveSortProgs{17}"
   Button "Button_85" at 864,635 size 256x28; TextOff 'Text'
      on Press: SetTag("Tag_1", 18)
      Visibility <- "DB939_Tool_alloc_HMI_SaveSortProgs{18}"
   Button "Button_86" at 864,662 size 256x28; TextOff 'Text'
      on Press: SetTag("Tag_1", 19)
      Visibility <- "DB939_Tool_alloc_HMI_SaveSortProgs{19}"
   Button "Button_87" at 864,689 size 256x28; TextOff 'Text'
      on Press: SetTag("Tag_1", 20)
      Visibility <- "DB939_Tool_alloc_HMI_SaveSortProgs{20}"
   Button "Button_88" at 118,149 size 306x41; TextOff 'Text'
      Visibility <- "DB939_Tool_alloc_HMI_Limit_allocation_list"
      on Press: SetTag("DB939_Tool_alloc_HMI_Selected_prog", 1)
   Button "Button_89" at 118,190 size 306x41; TextOff 'Text'
      on Press: SetTag("DB939_Tool_alloc_HMI_Selected_prog", 2)
      Visibility <- "DB939_Tool_alloc_HMI_Limit_allocation_list"
   Button "Button_90" at 118,230 size 306x41; TextOff 'Text'
      on Press: SetTag("DB939_Tool_alloc_HMI_Selected_prog", 3)
      Visibility <- "DB939_Tool_alloc_HMI_Limit_allocation_list"
   Button "Button_91" at 118,270 size 306x41; TextOff 'Text'
      on Press: SetTag("DB939_Tool_alloc_HMI_Selected_prog", 4)
      Visibility <- "DB939_Tool_alloc_HMI_Limit_allocation_list"
   Button "Button_92" at 118,310 size 306x41; TextOff 'Text'
      on Press: SetTag("DB939_Tool_alloc_HMI_Selected_prog", 5)
      Visibility <- "DB939_Tool_alloc_HMI_Limit_allocation_list"
   Button "Button_93" at 118,350 size 306x41; TextOff 'Text'
      on Press: SetTag("DB939_Tool_alloc_HMI_Selected_prog", 6)
      Visibility <- "DB939_Tool_alloc_HMI_Limit_allocation_list"
   Button "Button_94" at 118,390 size 306x41; TextOff 'Text'
      on Press: SetTag("DB939_Tool_alloc_HMI_Selected_prog", 7)
      Visibility <- "DB939_Tool_alloc_HMI_Limit_allocation_list"
   Button "Button_95" at 118,430 size 306x41; TextOff 'Text'
      on Press: SetTag("DB939_Tool_alloc_HMI_Selected_prog", 8)